   "PN_Mixinghead_Mixinghead{0}_DüseBypass{4}_Zeiten_Data_ÜberlappungD_B" : Real = PLC PN_Mixinghead.Mixinghead[0].DüseBypass[4].Zeiten.Data.ÜberlappungD_B AT %DB1006.DBD392, 1 s
      on ChangeValue: SetBit("PN_Mixinghead_Send"); SetBit("PN_Mixinghead_Mixinghead{0}_DüseBypass{4}_Zeiten_Request")
   "PN_Mixinghead_Mixinghead{0}_DüseBypass{4}_Zeiten_Data_ÜberlappungB_D" : Real = PLC PN_Mixinghead.Mixinghead[0].DüseBypass[4].Zeiten.Data.ÜberlappungB_D AT %DB1006.DBD396, 1 s
      on ChangeValue: SetBit("PN_Mixinghead_Send"); SetBit("PN_Mixinghead_Mixinghead{0}_DüseBypass{4}_Zeiten_Request")
   "PN_Mixinghead_Mixinghead{0}_DüseBypass{4}_Zeiten_Data_VerzögerungSchussstart" : Real = PLC PN_Mixinghead.Mixinghead[0].DüseBypass[4].Zeiten.Data.VerzögerungSchussstart AT %DB1006.DBD400, 1 s
      on ChangeValue: SetBit("PN_Mixinghead_Send"); SetBit("PN_Mixinghead_Mixinghead{0}_DüseBypass{4}_Zeiten_Request")
   "PN_Mixinghead_Mixinghead{0}_DüseBypass{4}_Zeiten_Data_VerzögerungSchussende" : Real = PLC PN_Mixinghead.Mixinghead[0].DüseBypass[4].Zeiten.Data.VerzögerungSchussende AT %DB1006.DBD404, 1 s
      on ChangeValue: SetBit("PN_Mixinghead_Send"); SetBit("PN_Mixinghead_Mixinghead{0}_DüseBypass{4}_Zeiten_Request")
   "PN_Mixinghead_Mixinghead{0}_DüseBypass{5}_Zeiten_Data_ÜberlappungD_B" : Real = PLC PN_Mixinghead.Mixinghead[0].DüseBypass[5].Zeiten.Data.ÜberlappungD_B AT %DB1006.DBD426, 1 s
      on ChangeValue: SetBit("PN_Mixinghead_Send"); SetBit("PN_Mixinghead_Mixinghead{0}_DüseBypass{5}_Zeiten_Request")
   "PN_Mixinghead_Mixinghead{0}_DüseBypass{5}_Zeiten_Data_ÜberlappungB_D" : Real = PLC PN_Mixinghead.Mixinghead[0].DüseBypass[5].Zeiten.Data.ÜberlappungB_D AT %DB1006.DBD430, 1 s
      on ChangeValue: SetBit("PN_Mixinghead_Send"); SetBit("PN_Mixinghead_Mixinghead{0}_DüseBypass{5}_Zeiten_Request")
   "PN_Mixinghead_Mixinghead{0}_DüseBypass{5}_Zeiten_Data_VerzögerungSchussstart" : Real = PLC PN_Mixinghead.Mixinghead[0].DüseBypass[5].Zeiten.Data.VerzögerungSchussstart AT %DB1006.DBD434, 1 s
      on ChangeValue: SetBit("PN_Mixinghead_Send"); SetBit("PN_Mixinghead_Mixinghead{0}_DüseBypass{5}_Zeiten_Request")
   "PN_Mixinghead_Mixinghead{0}_DüseBypass{5}_Zeiten_Data_VerzögerungSchussende" : Real = PLC PN_Mixinghead.Mixinghead[0].DüseBypass[5].Zeiten.Data.VerzögerungSchussende AT %DB1006.DBD438, 1 s
      on ChangeValue: SetBit("PN_Mixinghead_Send"); SetBit("PN_Mixinghead_Mixinghead{0}_DüseBypass{5}_Zeiten_Request")
   "PN_Mixinghead_Mixinghead{0}_DüseBypass{6}_Zeiten_Data_ÜberlappungD_B" : Real = PLC PN_Mixinghead.Mixinghead[0].DüseBypass[6].Zeiten.Data.ÜberlappungD_B AT %DB1006.DBD460, 1 s
      on ChangeValue: SetBit("PN_Mixinghead_Send"); SetBit("PN_Mixinghead_Mixinghead{0}_DüseBypass{6}_Zeiten_Request")
   "PN_Mixinghead_Mixinghead{0}_DüseBypass{6}_Zeiten_Data_ÜberlappungB_D" : Real = PLC PN_Mixinghead.Mixinghead[0].DüseBypass[6].Zeiten.Data.ÜberlappungB_D AT %DB1006.DBD464, 1 s
      on ChangeValue: SetBit("PN_Mixinghead_Send"); SetBit("PN_Mixinghead_Mixinghead{0}_DüseBypass{6}_Zeiten_Request")
   "PN_Mixinghead_Mixinghead{0}_DüseBypass{6}_Zeiten_Data_VerzögerungSchussstart" : Real = PLC PN_Mixinghead.Mixinghead[0].DüseBypass[6].Zeiten.Data.VerzögerungSchussstart AT %DB1006.DBD468, 1 s
      on ChangeValue: SetBit("PN_Mixinghead_Send"); SetBit("PN_Mixinghead_Mixinghead{0}_DüseBypass{6}_Zeiten_Request")
   "PN_Mixinghead_Mixinghead{0}_DüseBypass{6}_Zeiten_Data_VerzögerungSchussende" : Real = PLC PN_Mixinghead.Mixinghead[0].DüseBypass[6].Zeiten.Data.VerzögerungSchussende AT %DB1006.DBD472, 1 s
      on ChangeValue: SetBit("PN_Mixinghead_Send"); SetBit("PN_Mixinghead_Mixinghead{0}_DüseBypass{6}_Zeiten_Request")
   "PN_Error_Module{0}_AI{1}" : Int = PLC PN_Error.Module[0].AI[1] AT %DB1007.DBW112, 1 s
   "PN_Error_Module{0}_AI{2}" : Int = PLC PN_Error.Module[0].AI[2] AT %DB1007.DBW114, 1 s
   "PN_Error_Module{0}_AI{3}" : Int = PLC PN_Error.Module[0].AI[3] AT %DB1007.DBW116, 1 s
   "PN_Error_Module{0}_AI{4}" : Int = PLC PN_Error.Module[0].AI[4] AT %DB1007.DBW118, 1 s
   "PN_Error_Module{0}_AI{5}" : Int = PLC PN_Error.Module[0].AI[5] AT %DB1007.DBW120, 1 s
   "PN_Error_Module{0}_AI{6}" : Int = PLC PN_Error.Module[0].AI[6] AT %DB1007.DBW122, 1 s
   "PN_Error_Module{0}_AI{7}" : Int = PLC PN_Error.Module[0].AI[7] AT %DB1007.DBW124, 1 s
   "PN_Error_Module{0}_AI{8}" : Int = PLC PN_Error.Module[0].AI[8] AT %DB1007.DBW126, 1 s
   "PN_Error_Module{0}_AIr{1}" : Int = PLC PN_Error.Module[0].AIr[1] AT %DB1007.DBW128, 1 s
   "PN_Error_Module{0}_AIr{2}" : Int = PLC PN_Error.Module[0].AIr[2] AT %DB1007.DBW130, 1 s
   "PN_Error_Module{0}_AIr{3}" : Int = PLC PN_Error.Module[0].AIr[3] AT %DB1007.DBW132, 1 s
   "PN_Error_Module{0}_AIr{4}" : Int = PLC PN_Error.Module[0].AIr[4] AT %DB1007.DBW134, 1 s
   "PN_Error_Module{0}_AIr{5}" : Int = PLC PN_Error.Module[0].AIr[5] AT %DB1007.DBW136, 1 s
   "PN_Error_Module{0}_AIr{6}" : Int = PLC PN_Error.Module[0].AIr[6] AT %DB1007.DBW138, 1 s
   "PN_Error_Module{0}_AIr{7}" : Int = PLC PN_Error.Module[0].AIr[7] AT %DB1007.DBW140, 1 s
   "PN_Error_Module{0}_AIr{8}" : Int = PLC PN_Error.Module[0].AIr[8] AT %DB1007.DBW142, 1 s
   "PN_Error_Module{0}_DO_1" : DWord = PLC PN_Error.Module[0].DO_1 AT %DB1007.DBD104, 1 s
   "PN_Error_Module{0}_DO" : DWord = PLC PN_Error.Module[0].DO AT %DB1007.DBD108, 1 s
   "PN_AI_Module{0}_AI8_X14_0_Data_Data[3]_Bereichsobergrenze" : Int = PLC PN_AI.Module[0].AI8.X14_0.Data."Data[3]".Bereichsobergrenze AT %DB1002.DBW30, 1 s

HMI tags "Alarm"
   "Profibus_Alarm_DBW_16" : Int AT %DB820.DBW16, 1 s
      on ChangeValue: "RefreshAlarm"()
   "Profibus_Alarm_DBW_18" : Int AT %DB820.DBW18, 1 s
   "Profibus_Alarm_DBW_20" : Int AT %DB820.DBW20, 1 s
   "Profibus_Alarm_DBW_22" : Int AT %DB820.DBW22, 1 s
   "Profibus_Alarm_DBW_24" : Int AT %DB820.DBW24, 1 s
   "Profibus_Alarm_DBW_26" : Int AT %DB820.DBW26, 1 s
   "Profibus_Alarm_DBW_28" : Int AT %DB820.DBW28, 1 s
   "Profibus_Alarm_DBW_30" : Int AT %DB820.DBW30, 1 s
   "Machine_Alarm_DBW_58" : Int AT %DB820.DBW58, 1 s
      on ChangeValue: "RefreshAlarm"()
   "Machine_Alarm_DBW_60" : Int AT %DB820.DBW60, 1 s
      on ChangeValue: "RefreshAlarm"()
   "Machine_Alarm_DBW_62" : Int AT %DB820.DBW62, 1 s
      on ChangeValue: "RefreshAlarm"()
   "Machine_Alarm_DBW_64" : Int AT %DB820.DBW64, 1 s
   "Machine_Alarm_DBW_66" : Int AT %DB820.DBW66, 1 s
   "Interface_Container_DBW_520" : Int AT %DB822.DBW520, 1 s
   "Tank1_FeedPump_DBW_2" : Int AT %DB822.DBW2, 1 s
   "Tank2_FeedPump_DBW_4" : Int AT %DB822.DBW4, 1 s
   "Tank1_Agitator_DBW_28" : Int AT %DB822.DBW28, 1 s
   "Tank2_Agitator__DBW_30" : Int AT %DB822.DBW30, 1 s
   "Tank1_Filling_DBW_54" : Int AT %DB822.DBW54, 1 s
      on ChangeValue: "RefreshAlarm"()
   "Tank2_Filling_DBW_56" : Int AT %DB822.DBW56, 1 s
      on ChangeValue: "RefreshAlarm"()
   "Tank1_ControlerTemp_DBW_236" : Int AT %DB822.DBW236, 1 s
      on ChangeValue: "RefreshAlarm"()
   "Tank2_ControlerTemp_DBW_238" : Int AT %DB822.DBW238, 1 s
      on ChangeValue: "RefreshAlarm"()
   "Tank1_Pentan_DBW_496" : Int AT %DB822.DBW496, 1 s
   "Pump1_FeedPump_DBW_2" : Int AT %DB823.DBW2, 1 s
   "Pump1_EdgeFilter_DBW_28" : Int AT %DB823.DBW28, 1 s
   "Pump1_Component_DBW_56" : Int AT %DB823.DBW56, 1 s
      on ChangeValue: "RefreshAlarm"()
   "Pump1_Component_DBW_58" : Int AT %DB823.DBW58, 1 s
      on ChangeValue: "RefreshAlarm"()
   "Pump1_Flowrate_Record_DBW_106" : Int AT %DB823.DBW106, 1 s
   "Pump1_Pressure_Record_DBW_132" : Int AT %DB823.DBW132, 1 s
   "Pump1_Heatexchanger_DBW_210" : Int AT %DB823.DBW210, 1 s
   "Pump2_Component_DBW_60" : Int AT %DB823.DBW60, 1 s
      on ChangeValue: "RefreshAlarm"()
   "Pump2_Component_DBW_62" : Int AT %DB823.DBW62, 1 s
      on ChangeValue: "RefreshAlarm"()
   "Pump2_EdgeFilter_DBW_30" : Int AT %DB823.DBW30, 1 s
   "Pump2_FeedPump_DBW_4" : Int AT %DB823.DBW4, 1 s
   "Pump2_Flowrate_Record_DBW_108" : Int AT %DB823.DBW108, 1 s
   "Pump2_Heatexchanger_DBW_212" : Int AT %DB823.DBW212, 1 s
   "Pump2_Pressure_Record_DBW_134" : Int AT %DB823.DBW134, 1 s
   "Pump3_Component_DBW_64" : Int AT %DB823.DBW64, 1 s
   "Pump3_Component_DBW_66" : Int AT %DB823.DBW66, 1 s
   "Pump3_EdgeFilter_DBW_32" : Int AT %DB823.DBW32, 1 s
   "Pump3_FeedPump_DBW_6" : Int AT %DB823.DBW6, 1 s
   "Pump3_Flowrate_Record_DBW_110" : Int AT %DB823.DBW110, 1 s
   "Pump3_Heatexchanger_DBW_214" : Int AT %DB823.DBW214, 1 s
   "Pump3_Pressure_Record_DBW_136" : Int AT %DB823.DBW136, 1 s
   "Pump4_Component_DBW_68" : Int AT %DB823.DBW68, 1 s
   "Pump4_Component_DBW_70" : Int AT %DB823.DBW70, 1 s
   "Pump4_EdgeFilter_DBW_34" : Int AT %DB823.DBW34, 1 s
   "Pump4_FeedPump_DBW_8" : Int AT %DB823.DBW8, 1 s
   "Pump4_Flowrate_Record_DBW_112" : Int AT %DB823.DBW112, 1 s
   "Pump4_Heatexchanger_DBW_216" : Int AT %DB823.DBW216, 1 s
   "Pump4_Pressure_Record_DBW_138" : Int AT %DB823.DBW138, 1 s
   "Pump5_Component_DBW_72" : Int AT %DB823.DBW72, 1 s
   "Pump5_Component_DBW_74" : Int AT %DB823.DBW74, 1 s
   "Pump5_EdgeFilter_DBW_36" : Int AT %DB823.DBW36, 1 s
   "Pump5_FeedPump_DBW_10" : Int AT %DB823.DBW10, 1 s
   "Pump5_Flowrate_Record_DBW_114" : Int AT %DB823.DBW114, 1 s
   "Pump5_Heatexchanger_DBW_218" : Int AT %DB823.DBW218, 1 s
   "Pump5_Pressure_Record_DBW_140" : Int AT %DB823.DBW140, 1 s
   "Pump6_Component_DBW_76" : Int AT %DB823.DBW76, 1 s
   "Pump6_Component_DBW_78" : Int AT %DB823.DBW78, 1 s
   "Pump6_EdgeFilter_DBW_38" : Int AT %DB823.DBW38, 1 s
   "Pump6_FeedPump_DBW_12" : Int AT %DB823.DBW12, 1 s
   "Pump6_Flowrate_Record_DBW_116" : Int AT %DB823.DBW116, 1 s
   "Pump6_Heatexchanger_DBW_220" : Int AT %DB823.DBW220, 1 s
   "Pump6_Pressure_Record_DBW_142" : Int AT %DB823.DBW142, 1 s
   "Mixinghead_MHControl1_DBW_2" : Int AT %DB824.DBW2, 1 s
   "Mixinghead_MHControl2_DBW_4" : Int AT %DB824.DBW4, 1 s
   "Mixinghead_MHControl3_DBW_6" : Int AT %DB824.DBW6, 1 s
   "Mixinghead_MHControl4_DBW_8" : Int AT %DB824.DBW8, 1 s
   "Mixinghead_MHControl5_DBW_10" : Int AT %DB824.DBW10, 1 s
   "Mixinghead_MHControl6_DBW_12" : Int AT %DB824.DBW12, 1 s
   "Mixinghead_MHControl7_DBW_14" : Int AT %DB824.DBW14, 1 s
   "Mixinghead_MHControl8_DBW_16" : Int AT %DB824.DBW16, 1 s
   "Mixinghead_MHControl9_DBW_18" : Int AT %DB824.DBW18, 1 s
   "Mixinghead_MHControl10_DBW_20" : Int AT %DB824.DBW20, 1 s
   "Mixinghead_Cpiston1_DBW_34" : Int AT %DB824.DBW34, 1 s
      on ChangeValue: "RefreshAlarm"()
   "Mixinghead_Cpiston2_DBW_36" : Int AT %DB824.DBW36, 1 s
   "Mixinghead_Cpiston3_DBW_38" : Int AT %DB824.DBW38, 1 s
   "Mixinghead_Cpiston4_DBW_40" : Int AT %DB824.DBW40, 1 s
   "Mixinghead_Cpiston5_DBW_42" : Int AT %DB824.DBW42, 1 s
   "Mixinghead_Cpiston6_DBW_44" : Int AT %DB824.DBW44, 1 s
   "Mixinghead_Cpiston7_DBW_46" : Int AT %DB824.DBW46, 1 s
   "Mixinghead_Cpiston8_DBW_48" : Int AT %DB824.DBW48, 1 s
   "Mixinghead_Cpiston9_DBW_50" : Int AT %DB824.DBW50, 1 s
   "Mixinghead_Cpiston10_DBW_52" : Int AT %DB824.DBW52, 1 s
   "Mixinghead_Temperature_MH1_Con1_DBW70" : Int AT %DB824.DBW70, 1 s
      on ChangeValue: "RefreshAlarm"()
   "Mixinghead_Temperature_MH2_Con1_DBW72" : Int AT %DB824.DBW72, 1 s
   "Mixinghead_Temperature_MH3_Con1_DBW74" : Int AT %DB824.DBW74, 1 s
   "Mixinghead_Temperature_MH4_Con1_DBW76" : Int AT %DB824.DBW76, 1 s
   "Mixinghead_Temperature_MH5_Con1_DBW78" : Int AT %DB824.DBW78, 1 s
   "Mixinghead_Temperature_MH6_Con1_DBW80" : Int AT %DB824.DBW80, 1 s
   "Mixinghead_Temperature_MH7_Con1_DBW82" : Int AT %DB824.DBW82, 1 s
   "Mixinghead_Temperature_MH8_Con1_DBW84" : Int AT %DB824.DBW84, 1 s
   "Mixinghead_Temperature_MH9_Con1_DBW86" : Int AT %DB824.DBW86, 1 s
   "Mixinghead_Temperature_MH10_Con1_DBW88" : Int AT %DB824.DBW88, 1 s
   "Mixinghead_Temperature_MH1_Con2_DBW104" : Int AT %DB824.DBW104, 1 s
      on ChangeValue: "RefreshAlarm"()
   "Mixinghead_Temperature_MH2_Con2_DBW106" : Int AT %DB824.DBW106, 1 s
   "Mixinghead_Temperature_MH3_Con2_DBW108" : Int AT %DB824.DBW108, 1 s
   "Mixinghead_Temperature_MH4_Con2_DBW110" : Int AT %DB824.DBW110, 1 s
   "Mixinghead_Temperature_MH5_Con2_DBW112" : Int AT %DB824.DBW112, 1 s
   "Mixinghead_Temperature_MH6_Con2_DBW114" : Int AT %DB824.DBW114, 1 s
   "Mixinghead_Temperature_MH7_Con2_DBW116" : Int AT %DB824.DBW116, 1 s
   "Mixinghead_Temperature_MH8_Con2_DBW118" : Int AT %DB824.DBW118, 1 s
   "Mixinghead_Temperature_MH9_Con2_DBW120" : Int AT %DB824.DBW120, 1 s
   "Mixinghead_Temperature_MH10_Con2_DBW122" : Int AT %DB824.DBW122, 1 s
   "Mixinghead_Temperature_MH1_Con3_DBW138" : Int AT %DB824.DBW138, 1 s
      on ChangeValue: "RefreshAlarm"()
   "Mixinghead_Temperature_MH2_Con3_DBW140" : Int AT %DB824.DBW140, 1 s
   "Mixinghead_Temperature_MH3_Con3_DBW142" : Int AT %DB824.DBW142, 1 s
   "Mixinghead_Temperature_MH4_Con3_DBW144" : Int AT %DB824.DBW144, 1 s
   "Mixinghead_Temperature_MH5_Con3_DBW146" : Int AT %DB824.DBW146, 1 s
   "Mixinghead_Temperature_MH6_Con3_DBW148" : Int AT %DB824.DBW148, 1 s
   "Mixinghead_Temperature_MH7_Con3_DBW150" : Int AT %DB824.DBW150, 1 s
   "Mixinghead_Temperature_MH8_Con3_DBW152" : Int AT %DB824.DBW152, 1 s
   "Mixinghead_Temperature_MH9_Con3_DBW154" : Int AT %DB824.DBW154, 1 s
   "Mixinghead_Temperature_MH10_Con3_DBW156" : Int AT %DB824.DBW156, 1 s
   "Mixinghead_Temperature_MH1_Con4_DBW172" : Int AT %DB824.DBW172, 1 s
      on ChangeValue: "RefreshAlarm"()
   "Mixinghead_Temperature_MH2_Con4_DBW174" : Int AT %DB824.DBW174, 1 s
   "Mixinghead_Temperature_MH3_Con4_DBW176" : Int AT %DB824.DBW176, 1 s
   "Mixinghead_Temperature_MH4_Con4_DBW178" : Int AT %DB824.DBW178, 1 s
   "Mixinghead_Temperature_MH5_Con4_DBW180" : Int AT %DB824.DBW180, 1 s
   "Mixinghead_Temperature_MH6_Con4_DBW182" : Int AT %DB824.DBW182, 1 s
   "Mixinghead_Temperature_MH7_Con4_DBW184" : Int AT %DB824.DBW184, 1 s
   "Mixinghead_Temperature_MH8_Con4_DBW186" : Int AT %DB824.DBW186, 1 s
   "Mixinghead_Temperature_MH9_Con4_DBW188" : Int AT %DB824.DBW188, 1 s
   "Mixinghead_Temperature_MH10_Con4_DBW190" : Int AT %DB824.DBW190, 1 s
   "Mixinghead_Temperature_MH1_Con5_DBW206" : Int AT %DB824.DBW206, 1 s
      on ChangeValue: "RefreshAlarm"()
   "Mixinghead_Temperature_MH2_Con5_DBW208" : Int AT %DB824.DBW208, 1 s
   "Mixinghead_Temperature_MH3_Con5_DBW210" : Int AT %DB824.DBW210, 1 s
   "Mixinghead_Temperature_MH4_Con5_DBW212" : Int AT %DB824.DBW212, 1 s
   "Mixinghead_Temperature_MH5_Con5_DBW214" : Int AT %DB824.DBW214, 1 s
   "Mixinghead_Temperature_MH6_Con5_DBW216" : Int AT %DB824.DBW216, 1 s
   "Mixinghead_Temperature_MH7_Con5_DBW218" : Int AT %DB824.DBW218, 1 s
   "Mixinghead_Temperature_MH8_Con5_DBW220" : Int AT %DB824.DBW220, 1 s
   "Mixinghead_Temperature_MH9_Con5_DBW222" : Int AT %DB824.DBW222, 1 s
   "Mixinghead_Temperature_MH10_Con5_DBW224" : Int AT %DB824.DBW224, 1 s
   "Mixinghead_Temperature_MH1_Con6_DBW240" : Int AT %DB824.DBW240, 1 s
      on ChangeValue: "RefreshAlarm"()
   "Mixinghead_Temperature_MH2_Con6_DBW242" : Int AT %DB824.DBW242, 1 s
   "Mixinghead_Temperature_MH3_Con6_DBW244" : Int AT %DB824.DBW244, 1 s
   "Mixinghead_Temperature_MH4_Con6_DBW246" : Int AT %DB824.DBW246, 1 s
   "Mixinghead_Temperature_MH5_Con6_DBW248" : Int AT %DB824.DBW248, 1 s
   "Mixinghead_Temperature_MH6_Con6_DBW250" : Int AT %DB824.DBW250, 1 s
   "Mixinghead_Temperature_MH7_Con6_DBW252" : Int AT %DB824.DBW252, 1 s
   "Mixinghead_Temperature_MH8_Con6_DBW254" : Int AT %DB824.DBW254, 1 s
   "Mixinghead_Temperature_MH9_Con6_DBW256" : Int AT %DB824.DBW256, 1 s
   "Mixinghead_Temperature_MH10_Con6_DBW258" : Int AT %DB824.DBW258, 1 s
   "Mixinghead_Pressure_MH1_Con1_DBW274" : Int AT %DB824.DBW274, 1 s
   "Mixinghead_Pressure_MH2_Con1_DBW276" : Int AT %DB824.DBW276, 1 s
   "Mixinghead_Pressure_MH3_Con1_DBW278" : Int AT %DB824.DBW278, 1 s
   "Mixinghead_Pressure_MH4_Con1_DBW280" : Int AT %DB824.DBW280, 1 s
   "Mixinghead_Pressure_MH5_Con1_DBW282" : Int AT %DB824.DBW282, 1 s
   "Mixinghead_Pressure_MH6_Con1_DBW284" : Int AT %DB824.DBW284, 1 s
   "Mixinghead_Pressure_MH7_Con1_DBW286" : Int AT %DB824.DBW286, 1 s
   "Mixinghead_Pressure_MH8_Con1_DBW288" : Int AT %DB824.DBW288, 1 s
   "Mixinghead_Pressure_MH9_Con1_DBW290" : Int AT %DB824.DBW290, 1 s
   "Mixinghead_Pressure_MH10_Con1_DBW292" : Int AT %DB824.DBW292, 1 s
   "Mixinghead_Pressure_MH1_Con2_DBW308" : Int AT %DB824.DBW308, 1 s
   "Mixinghead_Pressure_MH2_Con2_DBW310" : Int AT %DB824.DBW310, 1 s
   "Mixinghead_Pressure_MH3_Con2_DBW312" : Int AT %DB824.DBW312, 1 s
   "Mixinghead_Pressure_MH4_Con2_DBW314" : Int AT %DB824.DBW314, 1 s
   "Mixinghead_Pressure_MH5_Con2_DBW316" : Int AT %DB824.DBW316, 1 s
   "Mixinghead_Pressure_MH6_Con2_DBW318" : Int AT %DB824.DBW318, 1 s
   "Mixinghead_Pressure_MH7_Con2_DBW320" : Int AT %DB824.DBW320, 1 s
   "Mixinghead_Pressure_MH8_Con2_DBW322" : Int AT %DB824.DBW322, 1 s
   "Mixinghead_Pressure_MH9_Con2_DBW324" : Int AT %DB824.DBW324, 1 s
   "Mixinghead_Pressure_MH10_Con2_DBW326" : Int AT %DB824.DBW326, 1 s
   "Mixinghead_Pressure_MH1_Con3_DBW342" : Int AT %DB824.DBW342, 1 s
   "Mixinghead_Pressure_MH2_Con3_DBW344" : Int AT %DB824.DBW344, 1 s
   "Mixinghead_Pressure_MH3_Con3_DBW346" : Int AT %DB824.DBW346, 1 s
   "Mixinghead_Pressure_MH4_Con3_DBW348" : Int AT %DB824.DBW348, 1 s
   "Mixinghead_Pressure_MH5_Con3_DBW350" : Int AT %DB824.DBW350, 1 s
   "Mixinghead_Pressure_MH6_Con3_DBW352" : Int AT %DB824.DBW352, 1 s
   "Mixinghead_Pressure_MH7_Con3_DBW354" : Int AT %DB824.DBW354, 1 s
   "Mixinghead_Pressure_MH8_Con3_DBW356" : Int AT %DB824.DBW356, 1 s
   "Mixinghead_Pressure_MH9_Con3_DBW358" : Int AT %DB824.DBW358, 1 s
   "Mixinghead_Pressure_MH10_Con3_DBW360" : Int AT %DB824.DBW360, 1 s
   "Mixinghead_Pressure_MH1_Con4_DBW376" : Int AT %DB824.DBW376, 1 s
   "Mixinghead_Pressure_MH2_Con4_DBW378" : Int AT %DB824.DBW378, 1 s
   "Mixinghead_Pressure_MH3_Con4_DBW380" : Int AT %DB824.DBW380, 1 s
   "Mixinghead_Pressure_MH4_Con4_DBW382" : Int AT %DB824.DBW382, 1 s
   "Mixinghead_Pressure_MH5_Con4_DBW384" : Int AT %DB824.DBW384, 1 s
   "Mixinghead_Pressure_MH6_Con4_DBW386" : Int AT %DB824.DBW386, 1 s
   "Mixinghead_Pressure_MH7_Con4_DBW388" : Int AT %DB824.DBW388, 1 s
   "Mixinghead_Pressure_MH8_Con4_DBW390" : Int AT %DB824.DBW390, 1 s
   "Mixinghead_Pressure_MH9_Con4_DBW392" : Int AT %DB824.DBW392, 1 s
   "Mixinghead_Pressure_MH10_Con4_DBW394" : Int AT %DB824.DBW394, 1 s
   "Mixinghead_Pressure_MH1_Con5_DBW410" : Int AT %DB824.DBW410, 1 s
   "Mixinghead_Pressure_MH2_Con5_DBW412" : Int AT %DB824.DBW412, 1 s
   "Mixinghead_Pressure_MH3_Con5_DBW414" : Int AT %DB824.DBW414, 1 s
   "Mixinghead_Pressure_MH4_Con5_DBW416" : Int AT %DB824.DBW416, 1 s
   "Mixinghead_Pressure_MH5_Con5_DBW418" : Int AT %DB824.DBW418, 1 s
   "Mixinghead_Pressure_MH6_Con5_DBW420" : Int AT %DB824.DBW420, 1 s
   "Mixinghead_Pressure_MH7_Con5_DBW422" : Int AT %DB824.DBW422, 1 s
   "Mixinghead_Pressure_MH8_Con5_DBW424" : Int AT %DB824.DBW424, 1 s
   "Mixinghead_Pressure_MH9_Con5_DBW426" : Int AT %DB824.DBW426, 1 s
   "Mixinghead_Pressure_MH10_Con5_DBW428" : Int AT %DB824.DBW428, 1 s
   "Mixinghead_Pressure_MH1_Con6_DBW444" : Int AT %DB824.DBW444, 1 s
   "Mixinghead_Pressure_MH2_Con6_DBW446" : Int AT %DB824.DBW446, 1 s
   "Mixinghead_Pressure_MH3_Con6_DBW448" : Int AT %DB824.DBW448, 1 s
   "Mixinghead_Pressure_MH4_Con6_DBW450" : Int AT %DB824.DBW450, 1 s
   "Mixinghead_Pressure_MH5_Con6_DBW452" : Int AT %DB824.DBW452, 1 s
   "Mixinghead_Pressure_MH6_Con6_DBW454" : Int AT %DB824.DBW454, 1 s
   "Mixinghead_Pressure_MH7_Con6_DBW456" : Int AT %DB824.DBW456, 1 s
   "Mixinghead_Pressure_MH8_Con6_DBW458" : Int AT %DB824.DBW458, 1 s
   "Mixinghead_Pressure_MH9_Con6_DBW460" : Int AT %DB824.DBW460, 1 s
   "Mixinghead_Pressure_MH10_Con6_DBW462" : Int AT %DB824.DBW462, 1 s
   "Mixinghead_Hydraulic_DBW2" : Int AT %DB821.DBW2, 1 s
   "Mixinghead_InertBlowout_MH1_DBW_546" : Int AT %DB824.DBW546, 1 s
   "Interface_MouldCarrier_1_DBW_0" : Int AT %DB825.DBW0, 1 s
   "Interface_MouldCarrier_2_DBW_2" : Int AT %DB825.DBW2, 1 s
   "Interface_MouldCarrier_3_DBW_4" : Int AT %DB825.DBW4, 1 s
   "Interface_MouldCarrier_4_DBW_6" : Int AT %DB825.DBW6, 1 s
   "Interface_MouldCarrier_5_DBW_8" : Int AT %DB825.DBW8, 1 s
   "Interface_MouldCarrier_6_DBW_10" : Int AT %DB825.DBW10, 1 s
   "Interface_MouldCarrier_7_DBW_12" : Int AT %DB825.DBW12, 1 s
   "Interface_MouldCarrier_8_DBW_14" : Int AT %DB825.DBW14, 1 s
   "Interface_MouldCarrier_9_DBW_16" : Int AT %DB825.DBW16, 1 s
   "Interface_MouldCarrier_10_DBW_18" : Int AT %DB825.DBW18, 1 s
   "Interface_External_1_DBW_32" : Int AT %DB825.DBW32, 1 s
   "Interface_Mould_Carrier_Emc_DBW_64" : Int AT %DB825.DBW64, 1 s
   "Error_Machine_SWU_DBW_0" : Int AT %DB829.DBW0, 1 s
   "Error_Machine_Pouring_DBW_4" : Int AT %DB829.DBW4, 1 s
      on ChangeValue: "RefreshAlarm"()
   "Error_Machine_Foaming_DBW_8" : Int AT %DB829.DBW8, 1 s
   "Machine_Filter_Alarm" : WString[30], internal
   "DosingPump_Filter_Alarm" : WString[10], internal
   "DB009_Faults_Fault_State_Grp_1_3_Exist" : Bool = PLC DB009_Faults.Fault_State_Grp_1_3_Exist AT %DB9.DBX1.7, 1 s
   "DB919_ShotResultMach_ShotResult_Ma{0}_General_PartWeight" : Real = PLC DB919_ShotResultMach.ShotResult_Ma[0].General.PartWeight AT %DB919.DBD48, 1 s
   "DB919_ShotResultMach_ShotResult_Ma{0}_General_FoamingTime" : Real = PLC DB919_ShotResultMach.ShotResult_Ma[0].General.FoamingTime AT %DB919.DBD52, 1 s
   "DB919_ShotResultMach_ShotResult_Ma{0}_General_StationNo" : Byte = PLC DB919_ShotResultMach.ShotResult_Ma[0].General.StationNo AT %DB919.DBB32, 1 s
   "DB919_ShotResultMach_ShotResult_Ma{0}_General_MH_No" : Byte = PLC DB919_ShotResultMach.ShotResult_Ma[0].General.MH_No AT %DB919.DBB34, 1 s
   "DB919_ShotResultMach_ShotResult_Ma{0}_General_ShotNo" : Int = PLC DB919_ShotResultMach.ShotResult_Ma[0].General.ShotNo AT %DB919.DBW16, 1 s
   "Foaming_Alarm" : Int, internal
   "DB919_ShotResultMach_ShotResult_Ma{0}_General_SendData" : Bool = PLC DB919_ShotResultMach.ShotResult_Ma[0].General.SendData AT %DB919.DBX0.0, 100 ms
      on ChangeValue: "FoamingAlarm"(); "RefreshAlarm"()
   "DB919_ShotResultMach_ShotResult_Ma{0}_Component_Comp{1}_Name" : String[20] = PLC DB919_ShotResultMach.ShotResult_Ma[0].Component.Comp[1].Name AT %DB919.DBX92.0, 1 s
   "DB919_ShotResultMach_ShotResult_Ma{0}_Component_Comp{1}_Flow" : Real = PLC DB919_ShotResultMach.ShotResult_Ma[0].Component.Comp[1].Flow AT %DB919.DBD120, 1 s
   "DB919_ShotResultMach_ShotResult_Ma{0}_Component_Comp{1}_PressureMH" : Real = PLC DB919_ShotResultMach.ShotResult_Ma[0].Component.Comp[1].PressureMH AT %DB919.DBD136, 1 s
   "DB919_ShotResultMach_ShotResult_Ma{0}_Component_Comp{1}_TemperatureMH" : Real = PLC DB919_ShotResultMach.ShotResult_Ma[0].Component.Comp[1].TemperatureMH AT %DB919.DBD152, 1 s
   "DB919_ShotResultMach_ShotResult_Ma{0}_Component_Comp{1}_Mixingratio" : Real = PLC DB919_ShotResultMach.ShotResult_Ma[0].Component.Comp[1].Mixingratio AT %DB919.DBD160, 1 s
   "DB919_ShotResultMach_ShotResult_Ma{0}_Component_Comp{2}_Name" : String[20] = PLC DB919_ShotResultMach.ShotResult_Ma[0].Component.Comp[2].Name AT %DB919.DBX168.0, 1 s
   "DB919_ShotResultMach_ShotResult_Ma{0}_Component_Comp{2}_Flow" : Real = PLC DB919_ShotResultMach.ShotResult_Ma[0].Component.Comp[2].Flow AT %DB919.DBD196, 1 s
   "DB919_ShotResultMach_ShotResult_Ma{0}_Component_Comp{2}_PressureMH" : Real = PLC DB919_ShotResultMach.ShotResult_Ma[0].Component.Comp[2].PressureMH AT %DB919.DBD212, 1 s
   "DB919_ShotResultMach_ShotResult_Ma{0}_Component_Comp{2}_TemperatureMH" : Real = PLC DB919_ShotResultMach.ShotResult_Ma[0].Component.Comp[2].TemperatureMH AT %DB919.DBD228, 1 s
   "DB919_ShotResultMach_ShotResult_Ma{0}_Component_Comp{2}_Mixingratio" : Real = PLC DB919_ShotResultMach.ShotResult_Ma[0].Component.Comp[2].Mixingratio AT %DB919.DBD236, 1 s
   "DB919_ShotResultMach_ShotResult_Ma{0}_Component_Comp{3}_Name" : String[20] = PLC DB919_ShotResultMach.ShotResult_Ma[0].Component.Comp[3].Name AT %DB919.DBX244.0, 1 s
   "DB919_ShotResultMach_ShotResult_Ma{0}_Component_Comp{3}_Flow" : Real = PLC DB919_ShotResultMach.ShotResult_Ma[0].Component.Comp[3].Flow AT %DB919.DBD272, 1 s
   "DB919_ShotResultMach_ShotResult_Ma{0}_Component_Comp{3}_PressureMH" : Real = PLC DB919_ShotResultMach.ShotResult_Ma[0].Component.Comp[3].PressureMH AT %DB919.DBD288, 1 s
   "DB919_ShotResultMach_ShotResult_Ma{0}_Component_Comp{3}_TemperatureMH" : Real = PLC DB919_ShotResultMach.ShotResult_Ma[0].Component.Comp[3].TemperatureMH AT %DB919.DBD304, 1 s
   "DB919_ShotResultMach_ShotResult_Ma{0}_Component_Comp{3}_Mixingratio" : Real = PLC DB919_ShotResultMach.ShotResult_Ma[0].Component.Comp[3].Mixingratio AT %DB919.DBD312, 1 s
   "DB919_ShotResultMach_ShotResult_Ma{0}_Component_Comp{4}_Name" : String[20] = PLC DB919_ShotResultMach.ShotResult_Ma[0].Component.Comp[4].Name AT %DB919.DBX320.0, 1 s
   "DB919_ShotResultMach_ShotResult_Ma{0}_Component_Comp{4}_Flow" : Real = PLC DB919_ShotResultMach.ShotResult_Ma[0].Component.Comp[4].Flow AT %DB919.DBD348, 1 s
   "DB919_ShotResultMach_ShotResult_Ma{0}_Component_Comp{4}_PressureMH" : Real = PLC DB919_ShotResultMach.ShotResult_Ma[0].Component.Comp[4].PressureMH AT %DB919.DBD364, 1 s
   "DB919_ShotResultMach_ShotResult_Ma{0}_Component_Comp{4}_TemperatureMH" : Real = PLC DB919_ShotResultMach.ShotResult_Ma[0].Component.Comp[4].TemperatureMH AT %DB919.DBD380, 1 s
   "DB919_ShotResultMach_ShotResult_Ma{0}_Component_Comp{4}_Mixingratio" : Real = PLC DB919_ShotResultMach.ShotResult_Ma[0].Component.Comp[4].Mixingratio AT %DB919.DBD388, 1 s
   "DB919_ShotResultMach_ShotResult_Ma{0}_Component_Comp{5}_Name" : String[20] = PLC DB919_ShotResultMach.ShotResult_Ma[0].Component.Comp[5].Name AT %DB919.DBX396.0, 1 s
   "DB919_ShotResultMach_ShotResult_Ma{0}_Component_Comp{5}_Flow" : Real = PLC DB919_ShotResultMach.ShotResult_Ma[0].Component.Comp[5].Flow AT %DB919.DBD424, 1 s
   "DB919_ShotResultMach_ShotResult_Ma{0}_Component_Comp{5}_PressureMH" : Real = PLC DB919_ShotResultMach.ShotResult_Ma[0].Component.Comp[5].PressureMH AT %DB919.DBD440, 1 s
   "DB919_ShotResultMach_ShotResult_Ma{0}_Component_Comp{5}_TemperatureMH" : Real = PLC DB919_ShotResultMach.ShotResult_Ma[0].Component.Comp[5].TemperatureMH AT %DB919.DBD456, 1 s
   "DB919_ShotResultMach_ShotResult_Ma{0}_Component_Comp{6}_Name" : String[20] = PLC DB919_ShotResultMach.ShotResult_Ma[0].Component.Comp[6].Name AT %DB919.DBX472.0, 1 s
   "DB919_ShotResultMach_ShotResult_Ma{0}_Component_Comp{6}_Flow" : Real = PLC DB919_ShotResultMach.ShotResult_Ma[0].Component.Comp[6].Flow AT %DB919.DBD500, 1 s
   "DB919_ShotResultMach_ShotResult_Ma{0}_Component_Comp{6}_PressureMH" : Real = PLC DB919_ShotResultMach.ShotResult_Ma[0].Component.Comp[6].PressureMH AT %DB919.DBD516, 1 s
   "DB919_ShotResultMach_ShotResult_Ma{0}_Component_Comp{6}_TemperatureMH" : Real = PLC DB919_ShotResultMach.ShotResult_Ma[0].Component.Comp[6].TemperatureMH AT %DB919.DBD532, 1 s
   "DB919_ShotResultMach_ShotResult_Ma{0}_Component_Comp{6}_Mixingratio" : Real = PLC DB919_ShotResultMach.ShotResult_Ma[0].Component.Comp[6].Mixingratio AT %DB919.DBD540, 1 s
   "DB919_ShotResultMach_ShotResult_Ma{0}_Component_Comp{7}_Name" : String[20] = PLC DB919_ShotResultMach.ShotResult_Ma[0].Component.Comp[7].Name AT %DB919.DBX548.0, 1 s
   "DB919_ShotResultMach_ShotResult_Ma{0}_Component_Comp{7}_Flow" : Real = PLC DB919_ShotResultMach.ShotResult_Ma[0].Component.Comp[7].Flow AT %DB919.DBD576, 1 s
   "DB919_ShotResultMach_ShotResult_Ma{0}_Component_Comp{7}_PressureMH" : Real = PLC DB919_ShotResultMach.ShotResult_Ma[0].Component.Comp[7].PressureMH AT %DB919.DBD592, 1 s
   "DB919_ShotResultMach_ShotResult_Ma{0}_Component_Comp{7}_TemperatureMH" : Real = PLC DB919_ShotResultMach.ShotResult_Ma[0].Component.Comp[7].TemperatureMH AT %DB919.DBD608, 1 s
   "DB919_ShotResultMach_ShotResult_Ma{0}_Component_Comp{7}_Mixingratio" : Real = PLC DB919_ShotResultMach.ShotResult_Ma[0].Component.Comp[7].Mixingratio AT %DB919.DBD616, 1 s
   "DB919_ShotResultMach_ShotResult_Ma{0}_Component_Comp{8}_Name" : String[20] = PLC DB919_ShotResultMach.ShotResult_Ma[0].Component.Comp[8].Name AT %DB919.DBX624.0, 1 s
   "DB919_ShotResultMach_ShotResult_Ma{0}_Component_Comp{8}_Flow" : Real = PLC DB919_ShotResultMach.ShotResult_Ma[0].Component.Comp[8].Flow AT %DB919.DBD652, 1 s
   "DB919_ShotResultMach_ShotResult_Ma{0}_Component_Comp{8}_PressureMH" : Real = PLC DB919_ShotResultMach.ShotResult_Ma[0].Component.Comp[8].PressureMH AT %DB919.DBD668, 1 s
   "DB919_ShotResultMach_ShotResult_Ma{0}_Component_Comp{8}_TemperatureMH" : Real = PLC DB919_ShotResultMach.ShotResult_Ma[0].Component.Comp[8].TemperatureMH AT %DB919.DBD684, 1 s
   "DB919_ShotResultMach_ShotResult_Ma{0}_Component_Comp{8}_Mixingratio" : Real = PLC DB919_ShotResultMach.ShotResult_Ma[0].Component.Comp[8].Mixingratio AT %DB919.DBD692, 1 s
   "DB919_ShotResultMach_ShotResult_Ma{0}_Component_Comp{9}_Name" : String[20] = PLC DB919_ShotResultMach.ShotResult_Ma[0].Component.Comp[9].Name AT %DB919.DBX700.0, 1 s
   "DB919_ShotResultMach_ShotResult_Ma{0}_Component_Comp{9}_Flow" : Real = PLC DB919_ShotResultMach.ShotResult_Ma[0].Component.Comp[9].Flow AT %DB919.DBD728, 1 s
   "DB919_ShotResultMach_ShotResult_Ma{0}_Component_Comp{9}_PressureMH" : Real = PLC DB919_ShotResultMach.ShotResult_Ma[0].Component.Comp[9].PressureMH AT %DB919.DBD744, 1 s
   "DB919_ShotResultMach_ShotResult_Ma{0}_Component_Comp{9}_TemperatureMH" : Real = PLC DB919_ShotResultMach.ShotResult_Ma[0].Component.Comp[9].TemperatureMH AT %DB919.DBD760, 1 s
   "DB919_ShotResultMach_ShotResult_Ma{0}_Component_Comp{9}_Mixingratio" : Real = PLC DB919_ShotResultMach.ShotResult_Ma[0].Component.Comp[9].Mixingratio AT %DB919.DBD768, 1 s
   "DB919_ShotResultMach_ShotResult_Ma{0}_Component_Comp{10}_Name" : String[20] = PLC DB919_ShotResultMach.ShotResult_Ma[0].Component.Comp[10].Name AT %DB919.DBX776.0, 1 s
   "DB919_ShotResultMach_ShotResult_Ma{0}_Component_Comp{10}_Flow" : Real = PLC DB919_ShotResultMach.ShotResult_Ma[0].Component.Comp[10].Flow AT %DB919.DBD804, 1 s
   "DB919_ShotResultMach_ShotResult_Ma{0}_Component_Comp{10}_PressureMH" : Real = PLC DB919_ShotResultMach.ShotResult_Ma[0].Component.Comp[10].PressureMH AT %DB919.DBD820, 1 s
   "DB919_ShotResultMach_ShotResult_Ma{0}_Component_Comp{10}_TemperatureMH" : Real = PLC DB919_ShotResultMach.ShotResult_Ma[0].Component.Comp[10].TemperatureMH AT %DB919.DBD836, 1 s
   "DB919_ShotResultMach_ShotResult_Ma{0}_Component_Comp{10}_Mixingratio" : Real = PLC DB919_ShotResultMach.ShotResult_Ma[0].Component.Comp[10].Mixingratio AT %DB919.DBD844, 1 s
   "DB919_ShotResultMach_ShotResult_Ma{0}_Component_Comp{11}_Name" : String[20] = PLC DB919_ShotResultMach.ShotResult_Ma[0].Component.Comp[11].Name AT %DB919.DBX852.0, 1 s
   "DB919_ShotResultMach_ShotResult_Ma{0}_Component_Comp{11}_Flow" : Real = PLC DB919_ShotResultMach.ShotResult_Ma[0].Component.Comp[11].Flow AT %DB919.DBD880, 1 s
   "DB919_ShotResultMach_ShotResult_Ma{0}_Component_Comp{11}_PressureMH" : Real = PLC DB919_ShotResultMach.ShotResult_Ma[0].Component.Comp[11].PressureMH AT %DB919.DBD896, 1 s
   "DB919_ShotResultMach_ShotResult_Ma{0}_Component_Comp{11}_TemperatureMH" : Real = PLC DB919_ShotResultMach.ShotResult_Ma[0].Component.Comp[11].TemperatureMH AT %DB919.DBD912, 1 s
   "DB919_ShotResultMach_ShotResult_Ma{0}_Component_Comp{11}_Mixingratio" : Real = PLC DB919_ShotResultMach.ShotResult_Ma[0].Component.Comp[11].Mixingratio AT %DB919.DBD920, 1 s
   "DB919_ShotResultMach_ShotResult_Ma{0}_Component_Comp{12}_Name" : String[20] = PLC DB919_ShotResultMach.ShotResult_Ma[0].Component.Comp[12].Name AT %DB919.DBX928.0, 1 s
   "DB919_ShotResultMach_ShotResult_Ma{0}_Component_Comp{12}_Flow" : Real = PLC DB919_ShotResultMach.ShotResult_Ma[0].Component.Comp[12].Flow AT %DB919.DBD956, 1 s
   "DB919_ShotResultMach_ShotResult_Ma{0}_Component_Comp{12}_PressureMH" : Real = PLC DB919_ShotResultMach.ShotResult_Ma[0].Component.Comp[12].PressureMH AT %DB919.DBD972, 1 s
   "DB919_ShotResultMach_ShotResult_Ma{0}_Component_Comp{12}_TemperatureMH" : Real = PLC DB919_ShotResultMach.ShotResult_Ma[0].Component.Comp[12].TemperatureMH AT %DB919.DBD988, 1 s
   "DB919_ShotResultMach_ShotResult_Ma{0}_Component_Comp{12}_Mixingratio" : Real = PLC DB919_ShotResultMach.ShotResult_Ma[0].Component.Comp[12].Mixingratio AT %DB919.DBD996, 1 s
   "DB919_ShotResultMach_ShotResult_Ma{0}_Component_Comp{5}_Mixingratio" : Real = PLC DB919_ShotResultMach.ShotResult_Ma[0].Component.Comp[5].Mixingratio AT %DB919.DBD464, 1 s
   "DB919_ShotResultMach_ShotResult_Ma{0}_Component_Comp{1}_ComponentActive" : Bool = PLC DB919_ShotResultMach.ShotResult_Ma[0].Component.Comp[1].ComponentActive AT %DB919.DBX114.0, 1 s
   "DB919_ShotResultMach_ShotResult_Ma{0}_Component_Comp{2}_ComponentActive" : Bool = PLC DB919_ShotResultMach.ShotResult_Ma[0].Component.Comp[2].ComponentActive AT %DB919.DBX190.0, 1 s
   "DB919_ShotResultMach_ShotResult_Ma{0}_Component_Comp{3}_ComponentActive" : Bool = PLC DB919_ShotResultMach.ShotResult_Ma[0].Component.Comp[3].ComponentActive AT %DB919.DBX266.0, 1 s
   "DB919_ShotResultMach_ShotResult_Ma{0}_Component_Comp{4}_ComponentActive" : Bool = PLC DB919_ShotResultMach.ShotResult_Ma[0].Component.Comp[4].ComponentActive AT %DB919.DBX342.0, 1 s
   "DB919_ShotResultMach_ShotResult_Ma{0}_Component_Comp{5}_ComponentActive" : Bool = PLC DB919_ShotResultMach.ShotResult_Ma[0].Component.Comp[5].ComponentActive AT %DB919.DBX418.0, 1 s
   "DB919_ShotResultMach_ShotResult_Ma{0}_Component_Comp{6}_ComponentActive" : Bool = PLC DB919_ShotResultMach.ShotResult_Ma[0].Component.Comp[6].ComponentActive AT %DB919.DBX494.0, 1 s
   "DB919_ShotResultMach_ShotResult_Ma{0}_Component_Comp{7}_ComponentActive" : Bool = PLC DB919_ShotResultMach.ShotResult_Ma[0].Component.Comp[7].ComponentActive AT %DB919.DBX570.0, 1 s
   "DB919_ShotResultMach_ShotResult_Ma{0}_Component_Comp{8}_ComponentActive" : Bool = PLC DB919_ShotResultMach.ShotResult_Ma[0].Component.Comp[8].ComponentActive AT %DB919.DBX646.0, 1 s

HMI tags "Service_PLC_Variabel"
   "DB1025_Service_State_Inputbyte" : Byte = PLC DB1025_Service.State.Inputbyte, 1 s
   "DB1025_Service_State_Outputbyte" : Byte = PLC DB1025_Service.State.Outputbyte, 1 s
   "DB1025_Service_Set_Inputbyte" : Word = PLC DB1025_Service.Set.Inputbyte, 1 s
   "DB1025_Service_Set_Outputbyte" : Word = PLC DB1025_Service.Set.Outputbyte, 1 s

HMI tags "System Setting"
   "TP-Bereichszeiger_Date_Time_ActTime_YEAR" : UInt = PLC "TP-Bereichszeiger".Date_Time.ActTime.YEAR AT %DB3.DBW44, 1 s
   "TP-Bereichszeiger_Date_Time_ActTime_MONTH" : USInt = PLC "TP-Bereichszeiger".Date_Time.ActTime.MONTH AT %DB3.DBB46, 1 s
   "TP-Bereichszeiger_Date_Time_ActTime_DAY" : USInt = PLC "TP-Bereichszeiger".Date_Time.ActTime.DAY AT %DB3.DBB47, 1 s
   "TP-Bereichszeiger_Date_Time_ActTime_WEEKDAY" : USInt = PLC "TP-Bereichszeiger".Date_Time.ActTime.WEEKDAY AT %DB3.DBB48, 1 s
   "TP-Bereichszeiger_Date_Time_ActTime_HOUR" : USInt = PLC "TP-Bereichszeiger".Date_Time.ActTime.HOUR AT %DB3.DBB49, 1 s
   "TP-Bereichszeiger_Date_Time_ActTime_MINUTE" : USInt = PLC "TP-Bereichszeiger".Date_Time.ActTime.MINUTE AT %DB3.DBB50, 1 s
   "TP-Bereichszeiger_Date_Time_ActTime_SECOND" : USInt = PLC "TP-Bereichszeiger".Date_Time.ActTime.SECOND AT %DB3.DBB51, 1 s
   "TP-Bereichszeiger_Date_Time_SetTime_YEAR" : UInt = PLC "TP-Bereichszeiger".Date_Time.SetTime.YEAR AT %DB3.DBW32, 1 s
   "TP-Bereichszeiger_Date_Time_SetTime_MONTH" : USInt = PLC "TP-Bereichszeiger".Date_Time.SetTime.MONTH AT %DB3.DBB34, 1 s
   "TP-Bereichszeiger_Date_Time_SetTime_DAY" : USInt = PLC "TP-Bereichszeiger".Date_Time.SetTime.DAY AT %DB3.DBB35, 1 s
   "TP-Bereichszeiger_Date_Time_SetTime_WEEKDAY" : USInt = PLC "TP-Bereichszeiger".Date_Time.SetTime.WEEKDAY AT %DB3.DBB36, 1 s
   "TP-Bereichszeiger_Date_Time_SetTime_HOUR" : USInt = PLC "TP-Bereichszeiger".Date_Time.SetTime.HOUR AT %DB3.DBB37, 1 s
   "TP-Bereichszeiger_Date_Time_SetTime_MINUTE" : USInt = PLC "TP-Bereichszeiger".Date_Time.SetTime.MINUTE AT %DB3.DBB38, 1 s
   "TP-Bereichszeiger_Date_Time_SetTime_SECOND" : USInt = PLC "TP-Bereichszeiger".Date_Time.SetTime.SECOND AT %DB3.DBB39, 1 s
   "TP-Bereichszeiger_Date_Time_Start_AG_Transfer" : Bool = PLC "TP-Bereichszeiger".Date_Time.Start_AG_Transfer AT %DB3.DBX30.0, 1 s
   "Operation Mode" : Int AT %DB619.DBW10, 1 s
   "DB619_State_MPart_Recirculation{1}_Intervall_Reduced" : Bool = PLC DB619_State_MPart.Recirculation[1].Intervall_Reduced AT %DB619.DBX44.4, 1 s
   "DB619_State_MPart_Recirculation{1}_Intervall_Lowpressure" : Bool = PLC DB619_State_MPart.Recirculation[1].Intervall_Lowpressure AT %DB619.DBX44.5, 1 s
   "DB619_State_MPart_Recirculation{1}_Intervall_Reduced_Pause" : Bool = PLC DB619_State_MPart.Recirculation[1].Intervall_Reduced_Pause AT %DB619.DBX44.6, 1 s
   "DB619_State_MPart_Recirculation{1}_Intervall_Lowpressure_Pause" : Bool = PLC DB619_State_MPart.Recirculation[1].Intervall_Lowpressure_Pause AT %DB619.DBX44.7, 1 s
   "DB619_State_MPart_Recirculation{1}_Highpressure" : Bool = PLC DB619_State_MPart.Recirculation[1].Highpressure AT %DB619.DBX42.4, 1 s
   "DB619_State_MPart_Recirculation{1}_Weekendswitching" : Bool = PLC DB619_State_MPart.Recirculation[1].Weekendswitching AT %DB619.DBX42.6, 1 s
   "DB619_State_MPart_Recirculation{1}_Lowpressure" : Bool = PLC DB619_State_MPart.Recirculation[1].Lowpressure AT %DB619.DBX42.2, 1 s
   "DB619_State_MPart_Recirculation{1}_Reduced" : Bool = PLC DB619_State_MPart.Recirculation[1].Reduced AT %DB619.DBX42.3, 1 s
   "DB619_State_MPart_Cycle{1}_running" : Bool = PLC DB619_State_MPart.Cycle[1].running AT %DB619.DBX222.1, 1 s
   "Print Function" : Bool AT %DB1.DBX0.0
   "TP-Bereichszeiger_Picturenumber_Bildnummer" : Int = PLC "TP-Bereichszeiger".Picturenumber.Bildnummer AT %DB3.DBW22, 1 s
   "TP-Bereichszeiger_Date_Time_ActTime" : DTL = PLC "TP-Bereichszeiger".Date_Time.ActTime AT %DB3.DBX44.0, 1 s
   "TP-Bereichszeiger_Koordinierungsbereich_Lebensbit" : Bool = PLC "TP-Bereichszeiger".Koordinierungsbereich.Lebensbit AT %DB3.DBX1.2, 500 ms
      on ChangeValue: "EndShift"()
   "TP-Bereichszeiger_Date_Time_SetTime" : DTL = PLC "TP-Bereichszeiger".Date_Time.SetTime AT %DB3.DBX32.0, 1 s
   "Computer_Name" : WString[20], internal
   "Ordner_Number" : WString[10], internal
   "Customer" : WString[45], internal
   "Additional_info_1" : WString[30], internal
   "Additional_info_2" : WString[30], internal
   "Additional_info_3" : WString[30], internal
   "Additional_info_5" : WString[30], internal
   "Additional_info_4" : WString[30], internal
   "Order_number" : WString[10], internal
   "Version" : WString[10], internal
   "Production_year" : WString[10], internal
   "Machine_number" : WString[10], internal
   "Wiring_diagram_number" : WString[10], internal

HMI tags "Create Part Counter"
   "Part_Counter_Name_1" : WString[20], internal
   "Part_Counter_Name_2" : WString[20], internal
   "Part_Counter_Name_3" : WString[20], internal
   "Part_Counter_Name_4" : WString[20], internal
   "Part_Counter_Name_5" : WString[20], internal
   "Part_Counter_Name_6" : WString[20], internal
   "Part_Counter_Name_7" : WString[20], internal
   "Part_Counter_Name_8" : WString[20], internal
   "Part_Counter_Name_9" : WString[20], internal
   "Part_Counter_Name_10" : WString[20], internal
   "Part_Counter_Name_11" : WString[20], internal
   "Part_Counter_Name_12" : WString[20], internal
   "Part_Counter_Name_13" : WString[20], internal
   "Part_Counter_Name_14" : WString[20], internal
   "Part_Counter_Name_15" : WString[20], internal
   "Part_Counter_Name_16" : WString[20], internal
   "Part_Counter_Name_17" : WString[20], internal
   "Part_Counter_Name_18" : WString[20], internal
   "Part_Counter_Name_19" : WString[20], internal
   "Part_Counter_Name_20" : WString[20], internal
   "Part_Counter_Name_21" : WString[20], internal
   "Part_Counter_Name_22" : WString[20], internal
   "Part_Counter_Name_23" : WString[20], internal
   "Part_Counter_Name_24" : WString[20], internal
   "Part_Counter_Name_25" : WString[20], internal
   "Part_Counter_Name_26" : WString[20], internal
   "Part_Counter_Name_27" : WString[20], internal
   "Part_Counter_Name_28" : WString[20], internal
   "Part_Counter_Name_29" : WString[20], internal
   "Part_Counter_Name_30" : WString[20], internal
   "Part_Counter_Name_31" : WString[20], internal
   "Part_Counter_Name_32" : WString[20], internal
   "Part_Counter_Name_33" : WString[20], internal
   "Part_Counter_Name_34" : WString[20], internal
   "Part_Counter_Name_35" : WString[20], internal
   "Part_Counter_Name_36" : WString[20], internal
   "Part_Counter_Name_37" : WString[20], internal
   "Part_Counter_Name_38" : WString[20], internal
   "Part_Counter_Name_39" : WString[20], internal
   "Part_Counter_Name_40" : WString[20], internal
   "Part_Counter_Name_41" : WString[20], internal
   "Part_Counter_Name_42" : WString[20], internal
   "Part_Counter_Name_43" : WString[20], internal
   "Part_Counter_Name_44" : WString[20], internal
   "Part_Counter_Name_45" : WString[20], internal
   "Part_Counter_Name_46" : WString[20], internal
   "Part_Counter_Name_47" : WString[20], internal
   "Part_Counter_Name_48" : WString[20], internal
   "Part_Counter_Name_49" : WString[20], internal
   "Part_Counter_Name_50" : WString[20], internal
   "Part_Counter_Name_51" : WString[20], internal
   "Part_Counter_Name_52" : WString[20], internal
   "Part_Counter_Name_53" : WString[20], internal
   "Part_Counter_Name_54" : WString[20], internal
   "Part_Counter_Name_55" : WString[20], internal
   "Part_Counter_Name_56" : WString[20], internal
   "Part_Counter_Name_57" : WString[20], internal
   "Part_Counter_Name_58" : WString[20], internal
   "Part_Counter_Name_59" : WString[20], internal
   "Part_Counter_Name_60" : WString[20], internal
   "Part_Counter_Name_61" : WString[20], internal
   "Part_Counter_Name_62" : WString[20], internal
   "Part_Counter_Name_63" : WString[20], internal
   "Part_Counter_Name_64" : WString[20], internal
   "Part_Counter_Name_65" : WString[20], internal
   "Part_Counter_Name_66" : WString[20], internal
   "Part_Counter_Name_67" : WString[20], internal
   "Part_Counter_Name_68" : WString[20], internal
   "Part_Counter_Name_69" : WString[20], internal
   "Part_Counter_Name_70" : WString[20], internal
   "Part_Counter_Name_71" : WString[20], internal
   "Part_Counter_Name_72" : WString[20], internal
   "Part_Counter_Name_73" : WString[20], internal
   "Part_Counter_Name_74" : WString[20], internal
   "Part_Counter_Name_75" : WString[20], internal
   "Part_Counter_Name_76" : WString[20], internal
   "Part_Counter_Name_77" : WString[20], internal
   "Part_Counter_Name_78" : WString[20], internal
   "Part_Counter_Name_79" : WString[20], internal
   "Part_Counter_Name_80" : WString[20], internal
   "Part_Counter_Name_81" : WString[20], internal
   "Part_Counter_Name_82" : WString[20], internal
   "Part_Counter_Name_83" : WString[20], internal
   "Part_Counter_Name_84" : WString[20], internal
   "Part_Counter_Name_85" : WString[20], internal
   "Part_Counter_Name_86" : WString[20], internal
   "Part_Counter_Name_87" : WString[20], internal
   "Part_Counter_Name_88" : WString[20], internal
   "Part_Counter_Name_89" : WString[20], internal
   "Part_Counter_Name_90" : WString[20], internal
   "Part_Counter_Name_91" : WString[20], internal
   "Part_Counter_Name_92" : WString[20], internal
   "Part_Counter_Name_93" : WString[20], internal
   "Part_Counter_Name_94" : WString[20], internal
   "Part_Counter_Name_95" : WString[20], internal
   "Part_Counter_Name_96" : WString[20], internal
   "Part_Counter_Name_97" : WString[20], internal
   "Part_Counter_Name_98" : WString[20], internal
   "Part_Counter_Name_99" : WString[20], internal
   "Part_Counter_Name_100" : WString[20], internal
   "Part_Counter_Name_101" : WString[20], internal
   "Part_Counter_Name_102" : WString[20], internal
   "Part_Counter_Name_103" : WString[20], internal
   "Part_Counter_Name_104" : WString[20], internal
   "Part_Counter_Name_105" : WString[20], internal
   "Part_Counter_Name_106" : WString[20], internal
   "Part_Counter_Name_107" : WString[20], internal
   "Part_Counter_Name_108" : WString[20], internal
   "Part_Counter_Name_109" : WString[20], internal
   "Part_Counter_Name_110" : WString[20], internal
   "Part_Counter_Name_111" : WString[20], internal
   "Part_Counter_Name_112" : WString[20], internal
   "Part_Counter_Name_113" : WString[20], internal
   "Part_Counter_Name_114" : WString[20], internal
   "Part_Counter_Name_115" : WString[20], internal
   "Part_Counter_Name_116" : WString[20], internal
   "Part_Counter_Name_117" : WString[20], internal
   "Part_Counter_Name_118" : WString[20], internal
   "Part_Counter_Name_119" : WString[20], internal
   "Part_Counter_Name_120" : WString[20], internal
   "Part_Counter_Coloum_1" : WString[10], internal
   "Part_Counter_Coloum_2" : WString[10], internal
   "Part_Counter_Coloum_3" : WString[10], internal
   "Part_Counter_Coloum_4" : WString[10], internal
   "Part_Counter_Coloum_5" : WString[10], internal
   "Part_Counter_Coloum_6" : WString[10], internal
   "Part_Counter_Coloum_7" : WString[10], internal
   "Part_Counter_Coloum_8" : WString[10], internal
   "Part_Counter_Coloum_9" : WString[10], internal
   "Part_Counter_Coloum_10" : WString[10], internal
   "Part_Counter_Coloum_11" : WString[10], internal
   "Part_Counter_Coloum_12" : WString[10], internal
   "Part_Counter_Coloum_13" : WString[10], internal
   "Part_Counter_Coloum_14" : WString[10], internal
   "Part_Counter_Coloum_15" : WString[10], internal
   "Part_Counter_Coloum_16" : WString[10], internal
   "Part_Counter_Coloum_17" : WString[10], internal
   "Part_Counter_Coloum_18" : WString[10], internal
   "Part_Counter_Coloum_19" : WString[10], internal
   "Part_Counter_Coloum_20" : WString[10], internal
   "Part_Counter_Coloum_21" : WString[10], internal
   "Part_Counter_Coloum_22" : WString[10], internal
   "Part_Counter_Coloum_23" : WString[10], internal
   "Part_Counter_Coloum_24" : WString[10], internal
   "Part_Counter_Coloum_25" : WString[10], internal
   "Part_Counter_Coloum_26" : WString[10], internal
   "Part_Counter_Coloum_27" : WString[10], internal
   "Part_Counter_Coloum_28" : WString[10], internal
   "Part_Counter_Coloum_29" : WString[10], internal
   "Part_Counter_Coloum_30" : WString[10], internal

